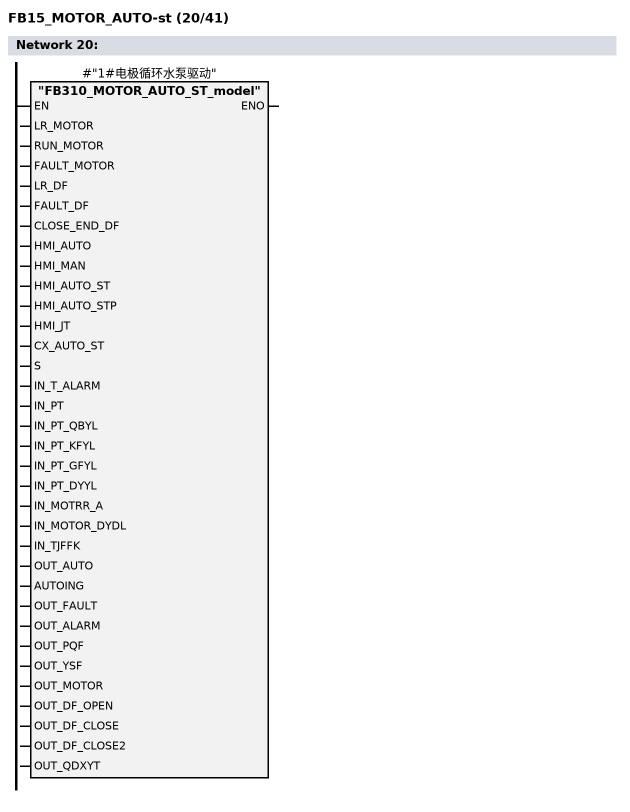
   RUNG wire#powerrail
      #"1#电极循环水泵驱动"(LR_MOTOR :=, RUN_MOTOR :=, FAULT_MOTOR :=, LR_DF :=, FAULT_DF :=, CLOSE_END_DF :=, HMI_AUTO :=, HMI_MAN :=, HMI_AUTO_ST :=, HMI_AUTO_STP :=, HMI_JT :=, CX_AUTO_ST :=, S :=, IN_T_ALARM :=, IN_PT :=, IN_PT_QBYL :=, IN_PT_KFYL :=, IN_PT_GFYL :=, IN_PT_DYYL :=, IN_MOTRR_A :=, IN_MOTOR_DYDL :=, IN_TJFFK :=, OUT_AUTO :=, AUTOING :=, OUT_FAULT :=, OUT_ALARM :=, OUT_PQF :=, OUT_YSF :=, OUT_MOTOR :=, OUT_DF_OPEN :=, OUT_DF_CLOSE :=, OUT_DF_CLOSE2 :=, OUT_QDXYT :=)
   END_RUNG
   // the same network as SCL:
   #"1#电极循环水泵驱动"();   // "FB310_MOTOR_AUTO_ST_model"
END_REGION

REGION Network 21
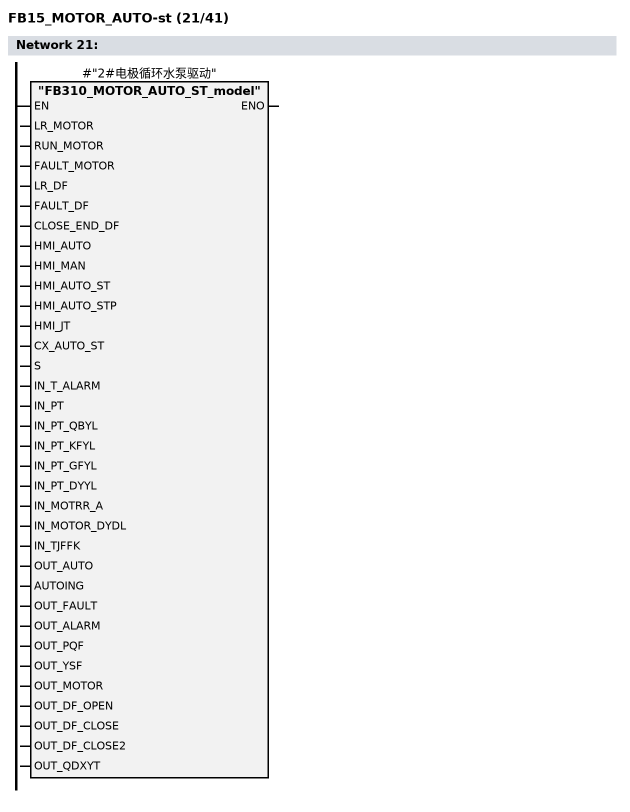
   RUNG wire#powerrail
      #"2#电极循环水泵驱动"(LR_MOTOR :=, RUN_MOTOR :=, FAULT_MOTOR :=, LR_DF :=, FAULT_DF :=, CLOSE_END_DF :=, HMI_AUTO :=, HMI_MAN :=, HMI_AUTO_ST :=, HMI_AUTO_STP :=, HMI_JT :=, CX_AUTO_ST :=, S :=, IN_T_ALARM :=, IN_PT :=, IN_PT_QBYL :=, IN_PT_KFYL :=, IN_PT_GFYL :=, IN_PT_DYYL :=, IN_MOTRR_A :=, IN_MOTOR_DYDL :=, IN_TJFFK :=, OUT_AUTO :=, AUTOING :=, OUT_FAULT :=, OUT_ALARM :=, OUT_PQF :=, OUT_YSF :=, OUT_MOTOR :=, OUT_DF_OPEN :=, OUT_DF_CLOSE :=, OUT_DF_CLOSE2 :=, OUT_QDXYT :=)
   END_RUNG
   // the same network as SCL:
   #"2#电极循环水泵驱动"();   // "FB310_MOTOR_AUTO_ST_model"
END_REGION

REGION Network 22
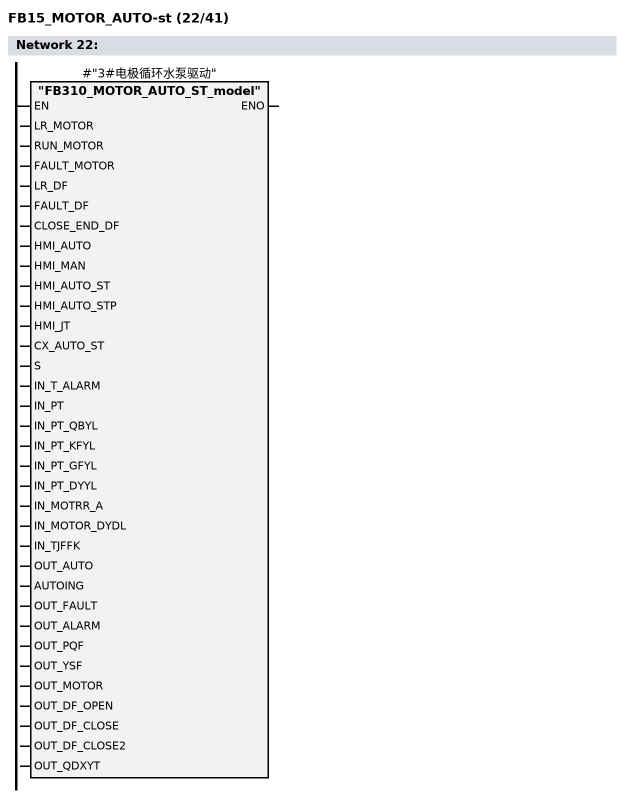
   RUNG wire#powerrail
      #"3#电极循环水泵驱动"(LR_MOTOR :=, RUN_MOTOR :=, FAULT_MOTOR :=, LR_DF :=, FAULT_DF :=, CLOSE_END_DF :=, HMI_AUTO :=, HMI_MAN :=, HMI_AUTO_ST :=, HMI_AUTO_STP :=, HMI_JT :=, CX_AUTO_ST :=, S :=, IN_T_ALARM :=, IN_PT :=, IN_PT_QBYL :=, IN_PT_KFYL :=, IN_PT_GFYL :=, IN_PT_DYYL :=, IN_MOTRR_A :=, IN_MOTOR_DYDL :=, IN_TJFFK :=, OUT_AUTO :=, AUTOING :=, OUT_FAULT :=, OUT_ALARM :=, OUT_PQF :=, OUT_YSF :=, OUT_MOTOR :=, OUT_DF_OPEN :=, OUT_DF_CLOSE :=, OUT_DF_CLOSE2 :=, OUT_QDXYT :=)
   END_RUNG
   // the same network as SCL:
   #"3#电极循环水泵驱动"();   // "FB310_MOTOR_AUTO_ST_model"
END_REGION

REGION Network 23
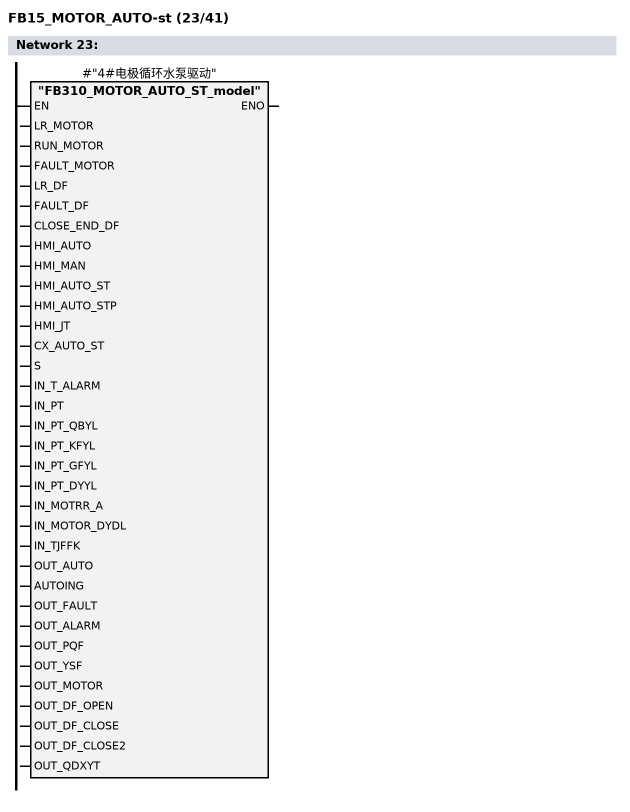
   RUNG wire#powerrail
      #"4#电极循环水泵驱动"(LR_MOTOR :=, RUN_MOTOR :=, FAULT_MOTOR :=, LR_DF :=, FAULT_DF :=, CLOSE_END_DF :=, HMI_AUTO :=, HMI_MAN :=, HMI_AUTO_ST :=, HMI_AUTO_STP :=, HMI_JT :=, CX_AUTO_ST :=, S :=, IN_T_ALARM :=, IN_PT :=, IN_PT_QBYL :=, IN_PT_KFYL :=, IN_PT_GFYL :=, IN_PT_DYYL :=, IN_MOTRR_A :=, IN_MOTOR_DYDL :=, IN_TJFFK :=, OUT_AUTO :=, AUTOING :=, OUT_FAULT :=, OUT_ALARM :=, OUT_PQF :=, OUT_YSF :=, OUT_MOTOR :=, OUT_DF_OPEN :=, OUT_DF_CLOSE :=, OUT_DF_CLOSE2 :=, OUT_QDXYT :=)
   END_RUNG
   // the same network as SCL:
   #"4#电极循环水泵驱动"();   // "FB310_MOTOR_AUTO_ST_model"
END_REGION

REGION Network 24
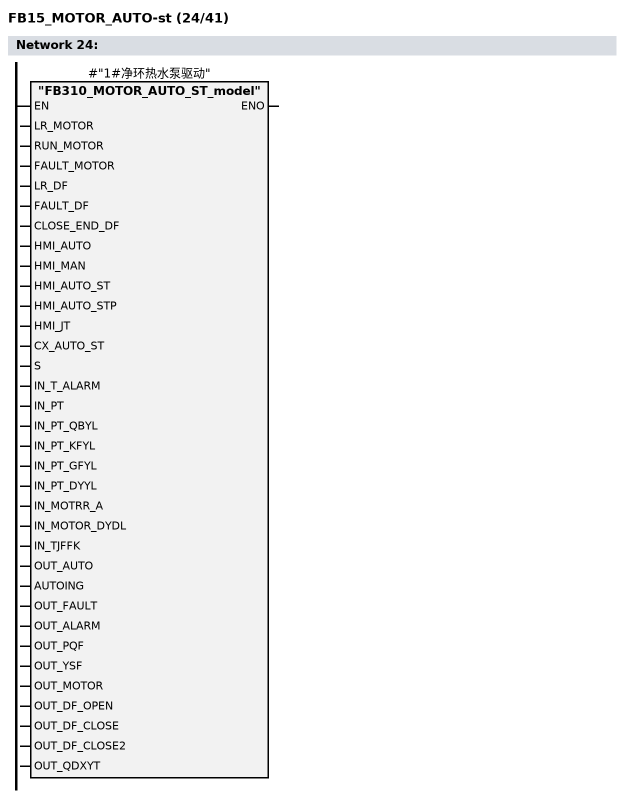
   RUNG wire#powerrail
      #"1#净环热水泵驱动"(LR_MOTOR :=, RUN_MOTOR :=, FAULT_MOTOR :=, LR_DF :=, FAULT_DF :=, CLOSE_END_DF :=, HMI_AUTO :=, HMI_MAN :=, HMI_AUTO_ST :=, HMI_AUTO_STP :=, HMI_JT :=, CX_AUTO_ST :=, S :=, IN_T_ALARM :=, IN_PT :=, IN_PT_QBYL :=, IN_PT_KFYL :=, IN_PT_GFYL :=, IN_PT_DYYL :=, IN_MOTRR_A :=, IN_MOTOR_DYDL :=, IN_TJFFK :=, OUT_AUTO :=, AUTOING :=, OUT_FAULT :=, OUT_ALARM :=, OUT_PQF :=, OUT_YSF :=, OUT_MOTOR :=, OUT_DF_OPEN :=, OUT_DF_CLOSE :=, OUT_DF_CLOSE2 :=, OUT_QDXYT :=)
   END_RUNG
   // the same network as SCL:
   #"1#净环热水泵驱动"();   // "FB310_MOTOR_AUTO_ST_model"
END_REGION

REGION Network 25
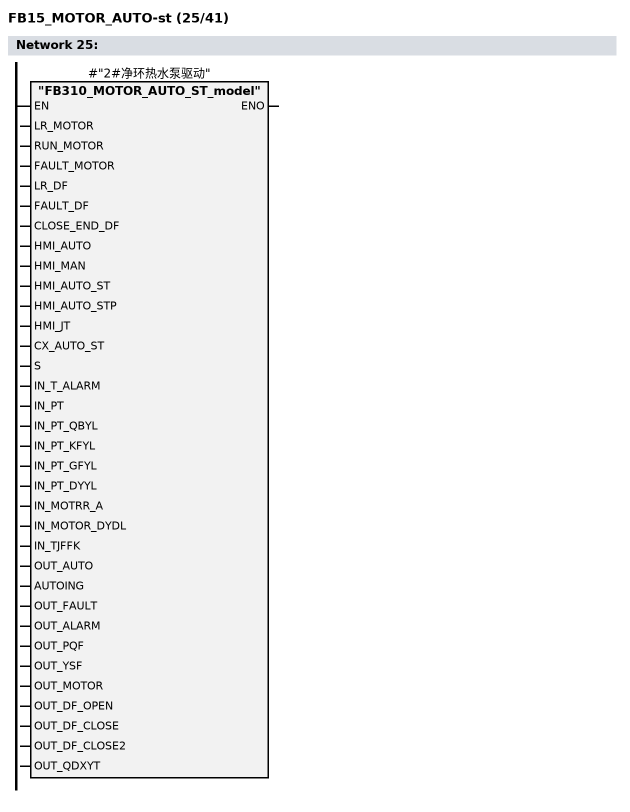
   RUNG wire#powerrail
      #"2#净环热水泵驱动"(LR_MOTOR :=, RUN_MOTOR :=, FAULT_MOTOR :=, LR_DF :=, FAULT_DF :=, CLOSE_END_DF :=, HMI_AUTO :=, HMI_MAN :=, HMI_AUTO_ST :=, HMI_AUTO_STP :=, HMI_JT :=, CX_AUTO_ST :=, S :=, IN_T_ALARM :=, IN_PT :=, IN_PT_QBYL :=, IN_PT_KFYL :=, IN_PT_GFYL :=, IN_PT_DYYL :=, IN_MOTRR_A :=, IN_MOTOR_DYDL :=, IN_TJFFK :=, OUT_AUTO :=, AUTOING :=, OUT_FAULT :=, OUT_ALARM :=, OUT_PQF :=, OUT_YSF :=, OUT_MOTOR :=, OUT_DF_OPEN :=, OUT_DF_CLOSE :=, OUT_DF_CLOSE2 :=, OUT_QDXYT :=)
   END_RUNG
   // the same network as SCL:
   #"2#净环热水泵驱动"();   // "FB310_MOTOR_AUTO_ST_model"
END_REGION

REGION Network 26
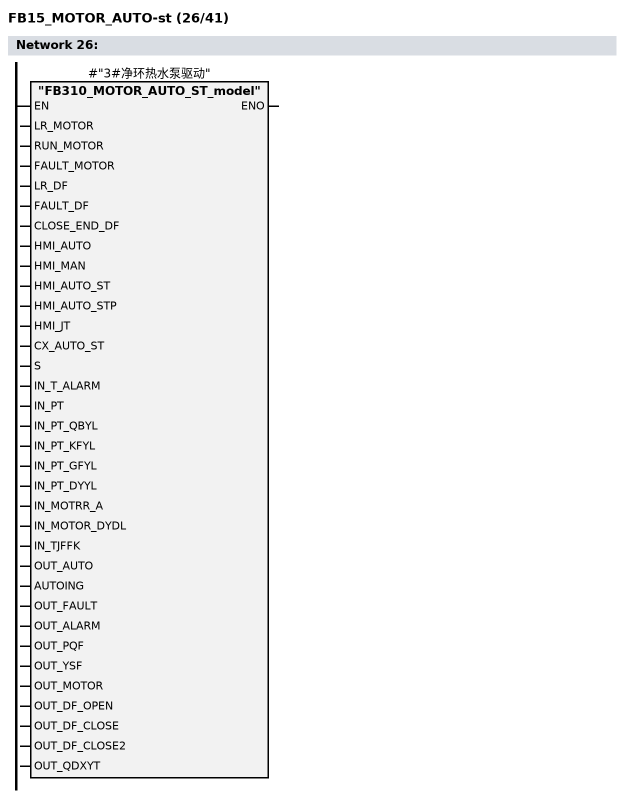
   RUNG wire#powerrail
      #"3#净环热水泵驱动"(LR_MOTOR :=, RUN_MOTOR :=, FAULT_MOTOR :=, LR_DF :=, FAULT_DF :=, CLOSE_END_DF :=, HMI_AUTO :=, HMI_MAN :=, HMI_AUTO_ST :=, HMI_AUTO_STP :=, HMI_JT :=, CX_AUTO_ST :=, S :=, IN_T_ALARM :=, IN_PT :=, IN_PT_QBYL :=, IN_PT_KFYL :=, IN_PT_GFYL :=, IN_PT_DYYL :=, IN_MOTRR_A :=, IN_MOTOR_DYDL :=, IN_TJFFK :=, OUT_AUTO :=, AUTOING :=, OUT_FAULT :=, OUT_ALARM :=, OUT_PQF :=, OUT_YSF :=, OUT_MOTOR :=, OUT_DF_OPEN :=, OUT_DF_CLOSE :=, OUT_DF_CLOSE2 :=, OUT_QDXYT :=)
   END_RUNG
   // the same network as SCL:
   #"3#净环热水泵驱动"();   // "FB310_MOTOR_AUTO_ST_model"
END_REGION

REGION Network 27
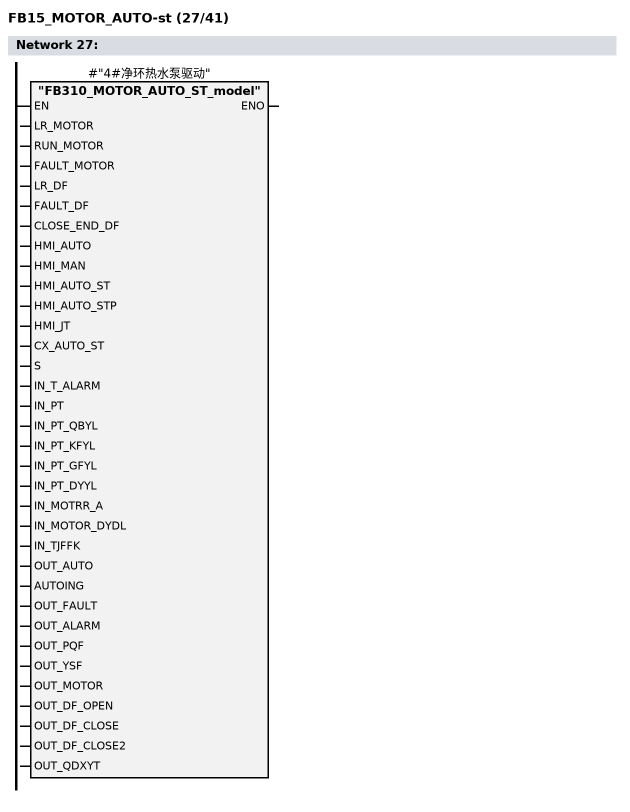
   RUNG wire#powerrail
      #"4#净环热水泵驱动"(LR_MOTOR :=, RUN_MOTOR :=, FAULT_MOTOR :=, LR_DF :=, FAULT_DF :=, CLOSE_END_DF :=, HMI_AUTO :=, HMI_MAN :=, HMI_AUTO_ST :=, HMI_AUTO_STP :=, HMI_JT :=, CX_AUTO_ST :=, S :=, IN_T_ALARM :=, IN_PT :=, IN_PT_QBYL :=, IN_PT_KFYL :=, IN_PT_GFYL :=, IN_PT_DYYL :=, IN_MOTRR_A :=, IN_MOTOR_DYDL :=, IN_TJFFK :=, OUT_AUTO :=, AUTOING :=, OUT_FAULT :=, OUT_ALARM :=, OUT_PQF :=, OUT_YSF :=, OUT_MOTOR :=, OUT_DF_OPEN :=, OUT_DF_CLOSE :=, OUT_DF_CLOSE2 :=, OUT_QDXYT :=)
   END_RUNG
   // the same network as SCL:
   #"4#净环热水泵驱动"();   // "FB310_MOTOR_AUTO_ST_model"
END_REGION

REGION Network 28
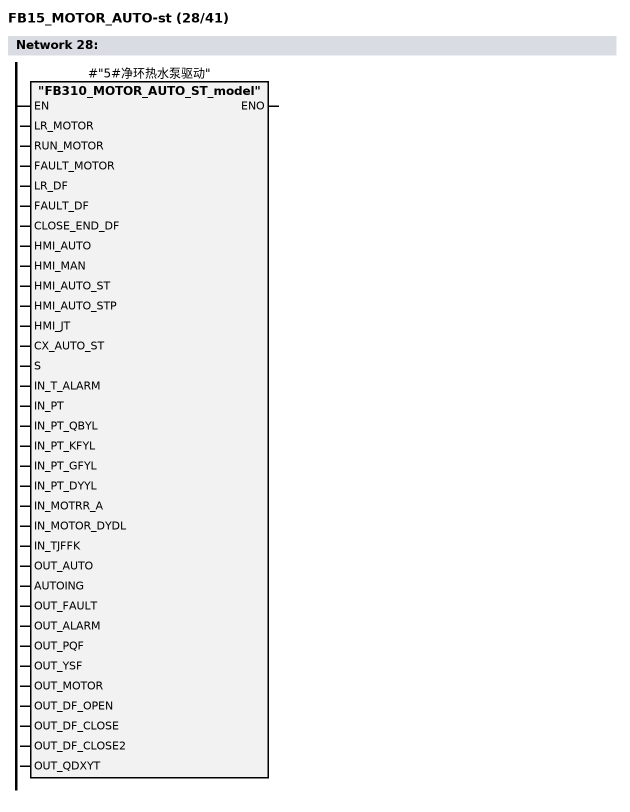
   RUNG wire#powerrail
      #"5#净环热水泵驱动"(LR_MOTOR :=, RUN_MOTOR :=, FAULT_MOTOR :=, LR_DF :=, FAULT_DF :=, CLOSE_END_DF :=, HMI_AUTO :=, HMI_MAN :=, HMI_AUTO_ST :=, HMI_AUTO_STP :=, HMI_JT :=, CX_AUTO_ST :=, S :=, IN_T_ALARM :=, IN_PT :=, IN_PT_QBYL :=, IN_PT_KFYL :=, IN_PT_GFYL :=, IN_PT_DYYL :=, IN_MOTRR_A :=, IN_MOTOR_DYDL :=, IN_TJFFK :=, OUT_AUTO :=, AUTOING :=, OUT_FAULT :=, OUT_ALARM :=, OUT_PQF :=, OUT_YSF :=, OUT_MOTOR :=, OUT_DF_OPEN :=, OUT_DF_CLOSE :=, OUT_DF_CLOSE2 :=, OUT_QDXYT :=)
   END_RUNG
   // the same network as SCL:
   #"5#净环热水泵驱动"();   // "FB310_MOTOR_AUTO_ST_model"
END_REGION

REGION Network 29
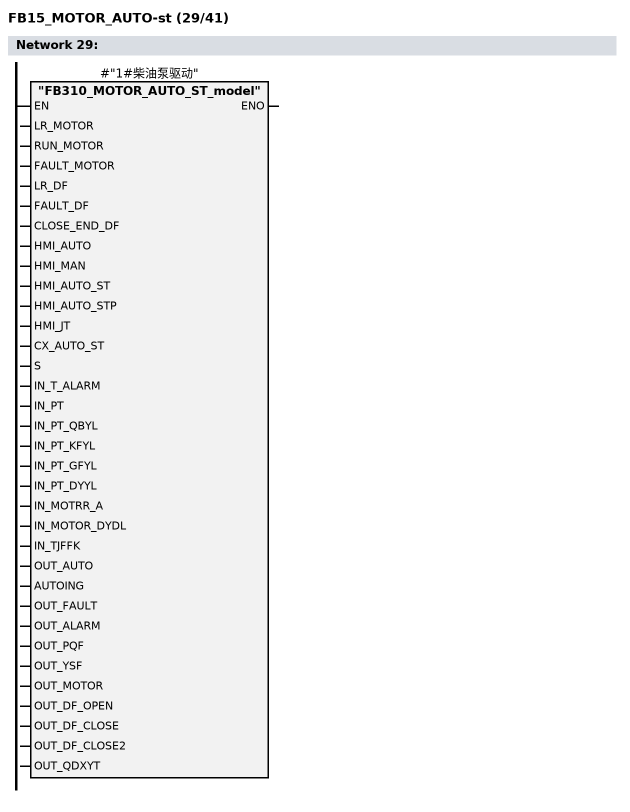
   RUNG wire#powerrail
      #"1#柴油泵驱动"(LR_MOTOR :=, RUN_MOTOR :=, FAULT_MOTOR :=, LR_DF :=, FAULT_DF :=, CLOSE_END_DF :=, HMI_AUTO :=, HMI_MAN :=, HMI_AUTO_ST :=, HMI_AUTO_STP :=, HMI_JT :=, CX_AUTO_ST :=, S :=, IN_T_ALARM :=, IN_PT :=, IN_PT_QBYL :=, IN_PT_KFYL :=, IN_PT_GFYL :=, IN_PT_DYYL :=, IN_MOTRR_A :=, IN_MOTOR_DYDL :=, IN_TJFFK :=, OUT_AUTO :=, AUTOING :=, OUT_FAULT :=, OUT_ALARM :=, OUT_PQF :=, OUT_YSF :=, OUT_MOTOR :=, OUT_DF_OPEN :=, OUT_DF_CLOSE :=, OUT_DF_CLOSE2 :=, OUT_QDXYT :=)
   END_RUNG
   // the same network as SCL:
   #"1#柴油泵驱动"();   // "FB310_MOTOR_AUTO_ST_model"
END_REGION

REGION Network 30
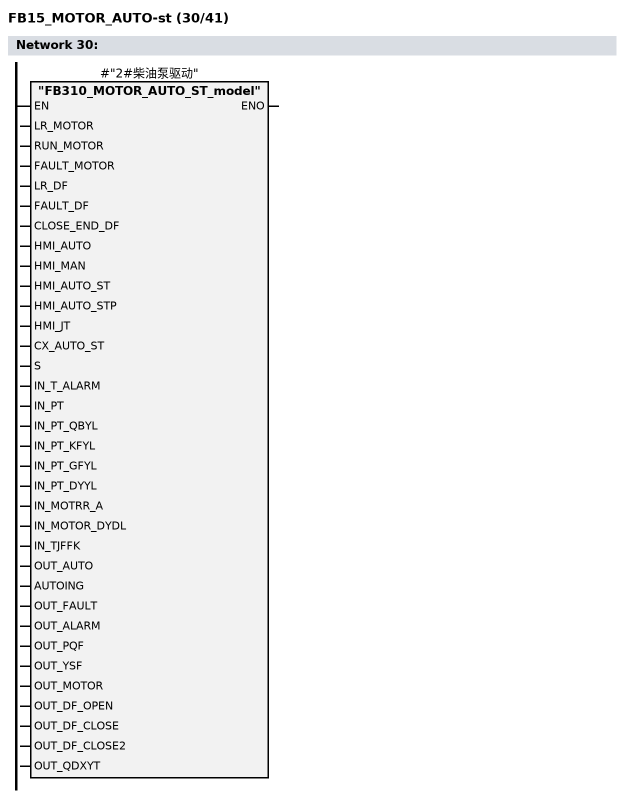
   RUNG wire#powerrail
      #"2#柴油泵驱动"(LR_MOTOR :=, RUN_MOTOR :=, FAULT_MOTOR :=, LR_DF :=, FAULT_DF :=, CLOSE_END_DF :=, HMI_AUTO :=, HMI_MAN :=, HMI_AUTO_ST :=, HMI_AUTO_STP :=, HMI_JT :=, CX_AUTO_ST :=, S :=, IN_T_ALARM :=, IN_PT :=, IN_PT_QBYL :=, IN_PT_KFYL :=, IN_PT_GFYL :=, IN_PT_DYYL :=, IN_MOTRR_A :=, IN_MOTOR_DYDL :=, IN_TJFFK :=, OUT_AUTO :=, AUTOING :=, OUT_FAULT :=, OUT_ALARM :=, OUT_PQF :=, OUT_YSF :=, OUT_MOTOR :=, OUT_DF_OPEN :=, OUT_DF_CLOSE :=, OUT_DF_CLOSE2 :=, OUT_QDXYT :=)
   END_RUNG
   // the same network as SCL:
   #"2#柴油泵驱动"();   // "FB310_MOTOR_AUTO_ST_model"
END_REGION

REGION Network 31
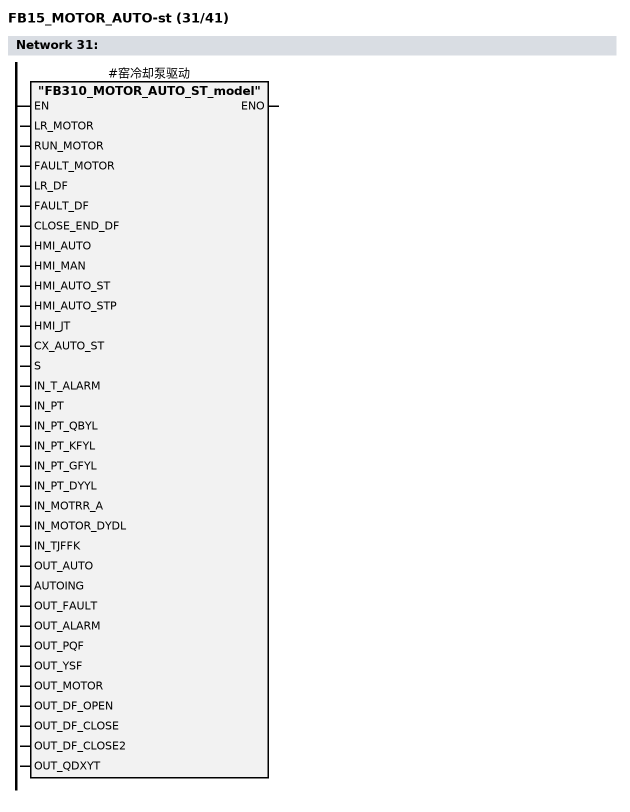
   RUNG wire#powerrail
      #窑冷却泵驱动(LR_MOTOR :=, RUN_MOTOR :=, FAULT_MOTOR :=, LR_DF :=, FAULT_DF :=, CLOSE_END_DF :=, HMI_AUTO :=, HMI_MAN :=, HMI_AUTO_ST :=, HMI_AUTO_STP :=, HMI_JT :=, CX_AUTO_ST :=, S :=, IN_T_ALARM :=, IN_PT :=, IN_PT_QBYL :=, IN_PT_KFYL :=, IN_PT_GFYL :=, IN_PT_DYYL :=, IN_MOTRR_A :=, IN_MOTOR_DYDL :=, IN_TJFFK :=, OUT_AUTO :=, AUTOING :=, OUT_FAULT :=, OUT_ALARM :=, OUT_PQF :=, OUT_YSF :=, OUT_MOTOR :=, OUT_DF_OPEN :=, OUT_DF_CLOSE :=, OUT_DF_CLOSE2 :=, OUT_QDXYT :=)
   END_RUNG
   // the same network as SCL:
   #窑冷却泵驱动();   // "FB310_MOTOR_AUTO_ST_model"
END_REGION

REGION Network 32
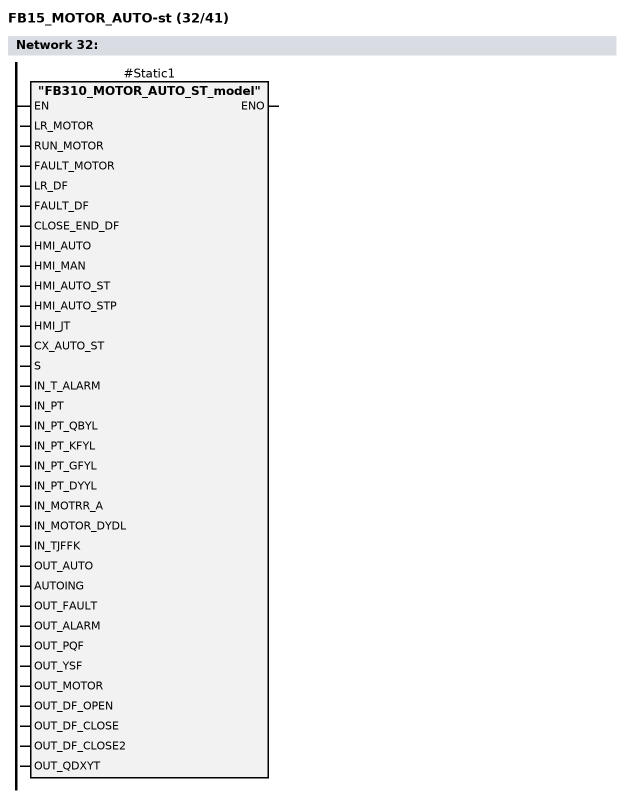
   RUNG wire#powerrail
      #Static1(LR_MOTOR :=, RUN_MOTOR :=, FAULT_MOTOR :=, LR_DF :=, FAULT_DF :=, CLOSE_END_DF :=, HMI_AUTO :=, HMI_MAN :=, HMI_AUTO_ST :=, HMI_AUTO_STP :=, HMI_JT :=, CX_AUTO_ST :=, S :=, IN_T_ALARM :=, IN_PT :=, IN_PT_QBYL :=, IN_PT_KFYL :=, IN_PT_GFYL :=, IN_PT_DYYL :=, IN_MOTRR_A :=, IN_MOTOR_DYDL :=, IN_TJFFK :=, OUT_AUTO :=, AUTOING :=, OUT_FAULT :=, OUT_ALARM :=, OUT_PQF :=, OUT_YSF :=, OUT_MOTOR :=, OUT_DF_OPEN :=, OUT_DF_CLOSE :=, OUT_DF_CLOSE2 :=, OUT_QDXYT :=)
   END_RUNG
   // the same network as SCL:
   #Static1();   // "FB310_MOTOR_AUTO_ST_model"
END_REGION

REGION Network 33
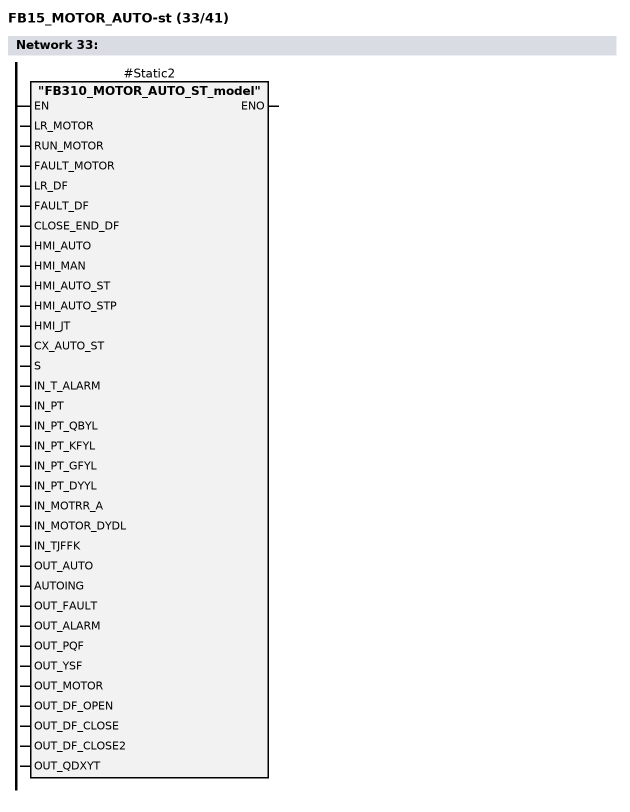
   RUNG wire#powerrail
      #Static2(LR_MOTOR :=, RUN_MOTOR :=, FAULT_MOTOR :=, LR_DF :=, FAULT_DF :=, CLOSE_END_DF :=, HMI_AUTO :=, HMI_MAN :=, HMI_AUTO_ST :=, HMI_AUTO_STP :=, HMI_JT :=, CX_AUTO_ST :=, S :=, IN_T_ALARM :=, IN_PT :=, IN_PT_QBYL :=, IN_PT_KFYL :=, IN_PT_GFYL :=, IN_PT_DYYL :=, IN_MOTRR_A :=, IN_MOTOR_DYDL :=, IN_TJFFK :=, OUT_AUTO :=, AUTOING :=, OUT_FAULT :=, OUT_ALARM :=, OUT_PQF :=, OUT_YSF :=, OUT_MOTOR :=, OUT_DF_OPEN :=, OUT_DF_CLOSE :=, OUT_DF_CLOSE2 :=, OUT_QDXYT :=)
   END_RUNG
   // the same network as SCL:
   #Static2();   // "FB310_MOTOR_AUTO_ST_model"
END_REGION

REGION Network 34
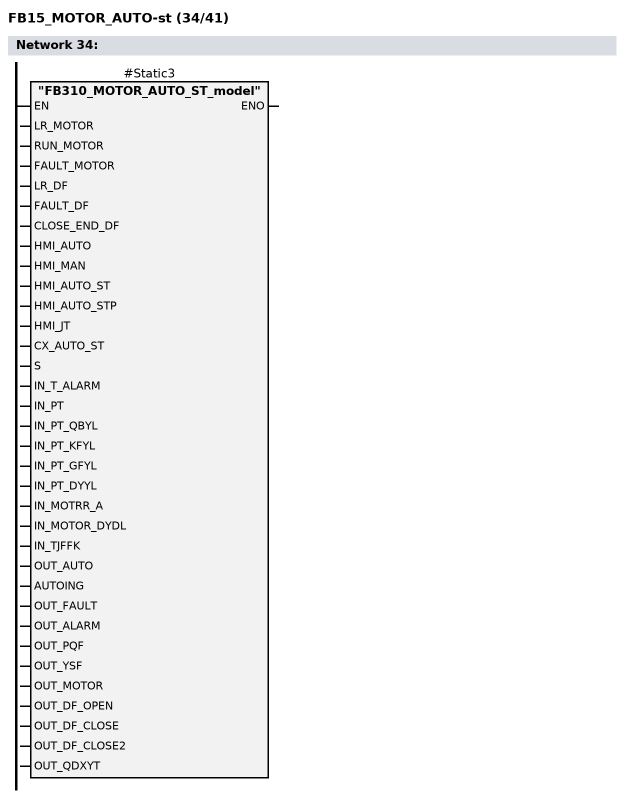
   RUNG wire#powerrail
      #Static3(LR_MOTOR :=, RUN_MOTOR :=, FAULT_MOTOR :=, LR_DF :=, FAULT_DF :=, CLOSE_END_DF :=, HMI_AUTO :=, HMI_MAN :=, HMI_AUTO_ST :=, HMI_AUTO_STP :=, HMI_JT :=, CX_AUTO_ST :=, S :=, IN_T_ALARM :=, IN_PT :=, IN_PT_QBYL :=, IN_PT_KFYL :=, IN_PT_GFYL :=, IN_PT_DYYL :=, IN_MOTRR_A :=, IN_MOTOR_DYDL :=, IN_TJFFK :=, OUT_AUTO :=, AUTOING :=, OUT_FAULT :=, OUT_ALARM :=, OUT_PQF :=, OUT_YSF :=, OUT_MOTOR :=, OUT_DF_OPEN :=, OUT_DF_CLOSE :=, OUT_DF_CLOSE2 :=, OUT_QDXYT :=)
   END_RUNG
   // the same network as SCL:
   #Static3();   // "FB310_MOTOR_AUTO_ST_model"
END_REGION

REGION Network 35
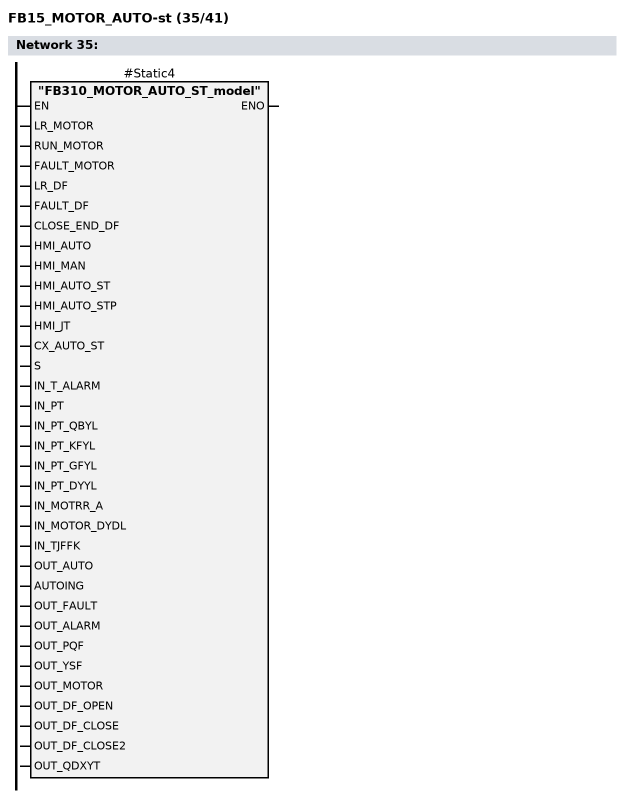
   RUNG wire#powerrail
      #Static4(LR_MOTOR :=, RUN_MOTOR :=, FAULT_MOTOR :=, LR_DF :=, FAULT_DF :=, CLOSE_END_DF :=, HMI_AUTO :=, HMI_MAN :=, HMI_AUTO_ST :=, HMI_AUTO_STP :=, HMI_JT :=, CX_AUTO_ST :=, S :=, IN_T_ALARM :=, IN_PT :=, IN_PT_QBYL :=, IN_PT_KFYL :=, IN_PT_GFYL :=, IN_PT_DYYL :=, IN_MOTRR_A :=, IN_MOTOR_DYDL :=, IN_TJFFK :=, OUT_AUTO :=, AUTOING :=, OUT_FAULT :=, OUT_ALARM :=, OUT_PQF :=, OUT_YSF :=, OUT_MOTOR :=, OUT_DF_OPEN :=, OUT_DF_CLOSE :=, OUT_DF_CLOSE2 :=, OUT_QDXYT :=)
   END_RUNG
   // the same network as SCL:
   #Static4();   // "FB310_MOTOR_AUTO_ST_model"
END_REGION

REGION Network 36
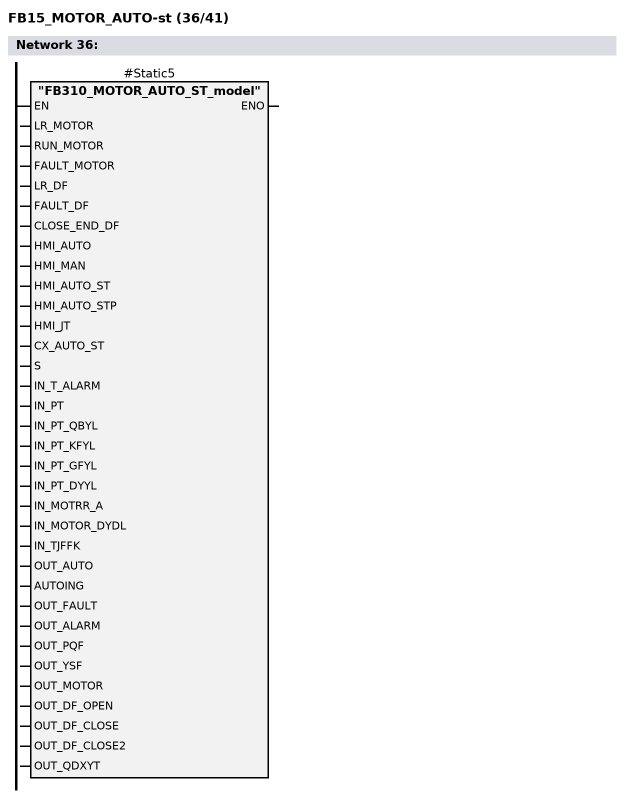
   RUNG wire#powerrail
      #Static5(LR_MOTOR :=, RUN_MOTOR :=, FAULT_MOTOR :=, LR_DF :=, FAULT_DF :=, CLOSE_END_DF :=, HMI_AUTO :=, HMI_MAN :=, HMI_AUTO_ST :=, HMI_AUTO_STP :=, HMI_JT :=, CX_AUTO_ST :=, S :=, IN_T_ALARM :=, IN_PT :=, IN_PT_QBYL :=, IN_PT_KFYL :=, IN_PT_GFYL :=, IN_PT_DYYL :=, IN_MOTRR_A :=, IN_MOTOR_DYDL :=, IN_TJFFK :=, OUT_AUTO :=, AUTOING :=, OUT_FAULT :=, OUT_ALARM :=, OUT_PQF :=, OUT_YSF :=, OUT_MOTOR :=, OUT_DF_OPEN :=, OUT_DF_CLOSE :=, OUT_DF_CLOSE2 :=, OUT_QDXYT :=)
   END_RUNG
   // the same network as SCL:
   #Static5();   // "FB310_MOTOR_AUTO_ST_model"
END_REGION

REGION Network 37
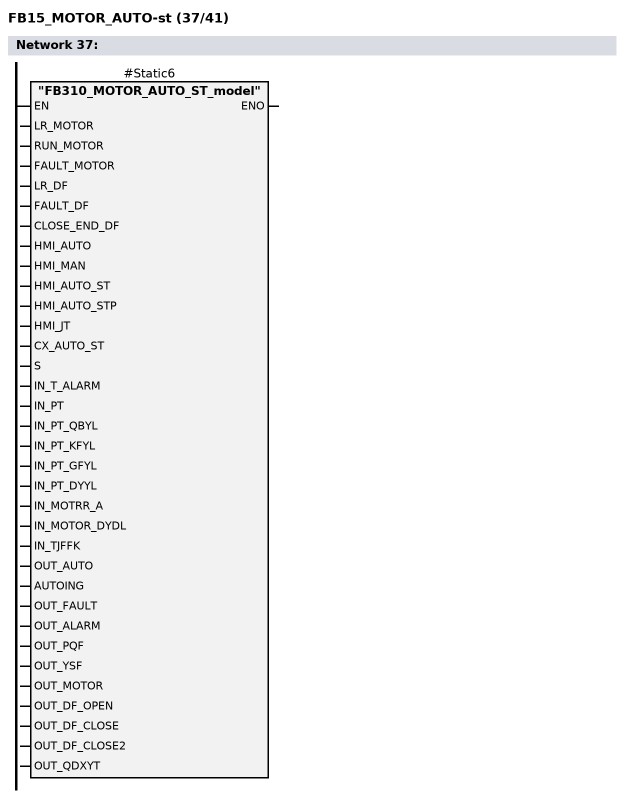
   RUNG wire#powerrail
      #Static6(LR_MOTOR :=, RUN_MOTOR :=, FAULT_MOTOR :=, LR_DF :=, FAULT_DF :=, CLOSE_END_DF :=, HMI_AUTO :=, HMI_MAN :=, HMI_AUTO_ST :=, HMI_AUTO_STP :=, HMI_JT :=, CX_AUTO_ST :=, S :=, IN_T_ALARM :=, IN_PT :=, IN_PT_QBYL :=, IN_PT_KFYL :=, IN_PT_GFYL :=, IN_PT_DYYL :=, IN_MOTRR_A :=, IN_MOTOR_DYDL :=, IN_TJFFK :=, OUT_AUTO :=, AUTOING :=, OUT_FAULT :=, OUT_ALARM :=, OUT_PQF :=, OUT_YSF :=, OUT_MOTOR :=, OUT_DF_OPEN :=, OUT_DF_CLOSE :=, OUT_DF_CLOSE2 :=, OUT_QDXYT :=)
   END_RUNG
   // the same network as SCL:
   #Static6();   // "FB310_MOTOR_AUTO_ST_model"
END_REGION

REGION Network 38
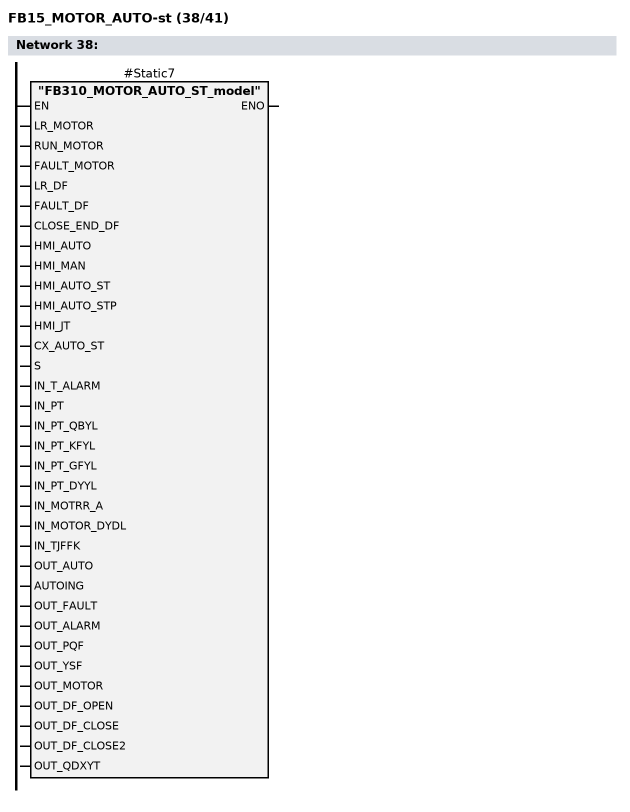
   RUNG wire#powerrail
      #Static7(LR_MOTOR :=, RUN_MOTOR :=, FAULT_MOTOR :=, LR_DF :=, FAULT_DF :=, CLOSE_END_DF :=, HMI_AUTO :=, HMI_MAN :=, HMI_AUTO_ST :=, HMI_AUTO_STP :=, HMI_JT :=, CX_AUTO_ST :=, S :=, IN_T_ALARM :=, IN_PT :=, IN_PT_QBYL :=, IN_PT_KFYL :=, IN_PT_GFYL :=, IN_PT_DYYL :=, IN_MOTRR_A :=, IN_MOTOR_DYDL :=, IN_TJFFK :=, OUT_AUTO :=, AUTOING :=, OUT_FAULT :=, OUT_ALARM :=, OUT_PQF :=, OUT_YSF :=, OUT_MOTOR :=, OUT_DF_OPEN :=, OUT_DF_CLOSE :=, OUT_DF_CLOSE2 :=, OUT_QDXYT :=)
   END_RUNG
   // the same network as SCL:
   #Static7();   // "FB310_MOTOR_AUTO_ST_model"
END_REGION

REGION Network 39
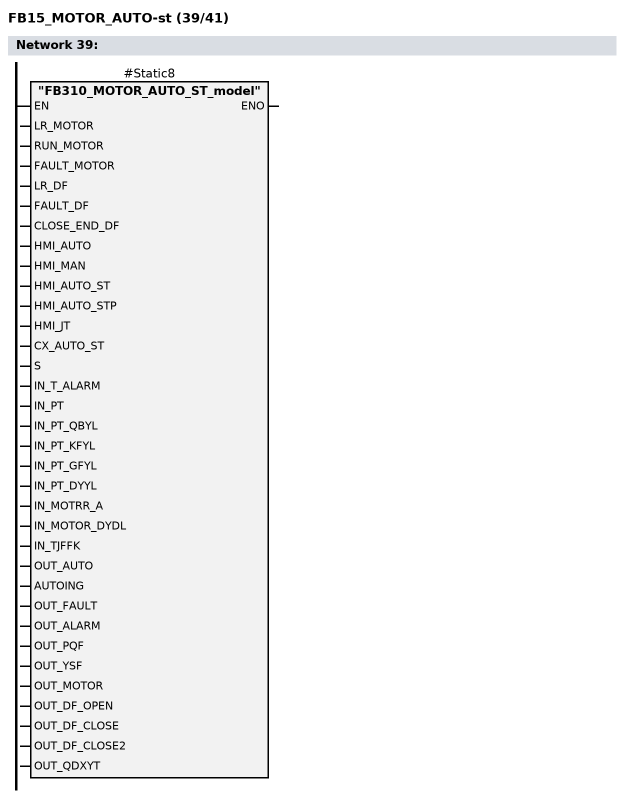
   RUNG wire#powerrail
      #Static8(LR_MOTOR :=, RUN_MOTOR :=, FAULT_MOTOR :=, LR_DF :=, FAULT_DF :=, CLOSE_END_DF :=, HMI_AUTO :=, HMI_MAN :=, HMI_AUTO_ST :=, HMI_AUTO_STP :=, HMI_JT :=, CX_AUTO_ST :=, S :=, IN_T_ALARM :=, IN_PT :=, IN_PT_QBYL :=, IN_PT_KFYL :=, IN_PT_GFYL :=, IN_PT_DYYL :=, IN_MOTRR_A :=, IN_MOTOR_DYDL :=, IN_TJFFK :=, OUT_AUTO :=, AUTOING :=, OUT_FAULT :=, OUT_ALARM :=, OUT_PQF :=, OUT_YSF :=, OUT_MOTOR :=, OUT_DF_OPEN :=, OUT_DF_CLOSE :=, OUT_DF_CLOSE2 :=, OUT_QDXYT :=)
   END_RUNG
   // the same network as SCL:
   #Static8();   // "FB310_MOTOR_AUTO_ST_model"
END_REGION

REGION Network 40
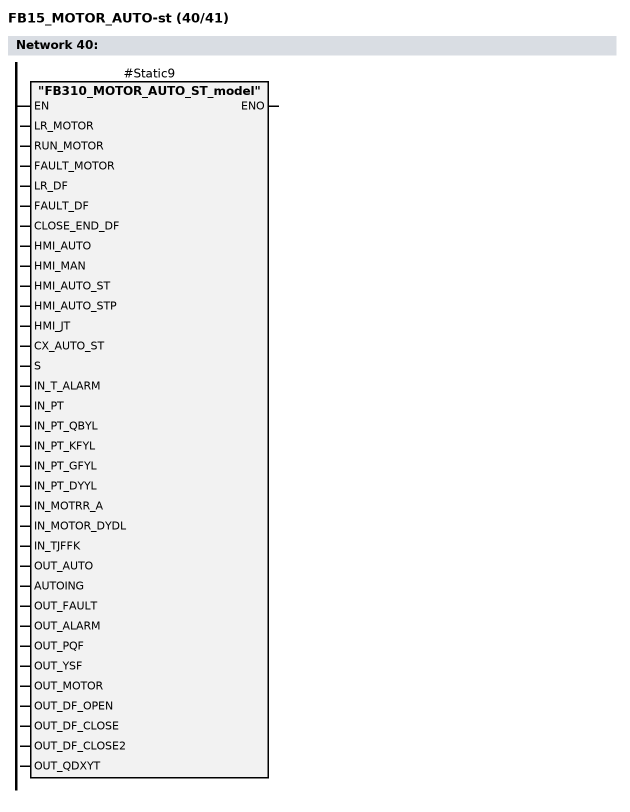
   RUNG wire#powerrail
      #Static9(LR_MOTOR :=, RUN_MOTOR :=, FAULT_MOTOR :=, LR_DF :=, FAULT_DF :=, CLOSE_END_DF :=, HMI_AUTO :=, HMI_MAN :=, HMI_AUTO_ST :=, HMI_AUTO_STP :=, HMI_JT :=, CX_AUTO_ST :=, S :=, IN_T_ALARM :=, IN_PT :=, IN_PT_QBYL :=, IN_PT_KFYL :=, IN_PT_GFYL :=, IN_PT_DYYL :=, IN_MOTRR_A :=, IN_MOTOR_DYDL :=, IN_TJFFK :=, OUT_AUTO :=, AUTOING :=, OUT_FAULT :=, OUT_ALARM :=, OUT_PQF :=, OUT_YSF :=, OUT_MOTOR :=, OUT_DF_OPEN :=, OUT_DF_CLOSE :=, OUT_DF_CLOSE2 :=, OUT_QDXYT :=)
   END_RUNG
   // the same network as SCL:
   #Static9();   // "FB310_MOTOR_AUTO_ST_model"
END_REGION

REGION Network 41
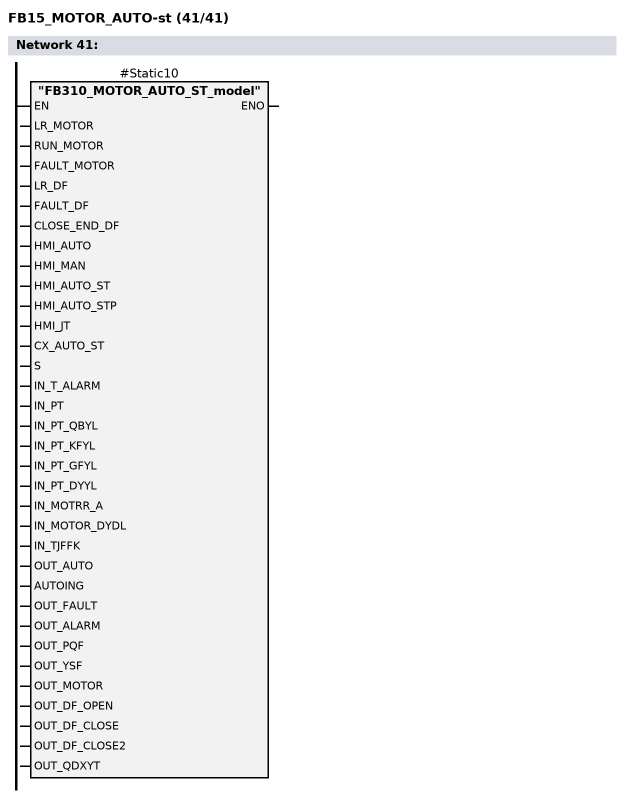
   RUNG wire#powerrail
      #Static10(LR_MOTOR :=, RUN_MOTOR :=, FAULT_MOTOR :=, LR_DF :=, FAULT_DF :=, CLOSE_END_DF :=, HMI_AUTO :=, HMI_MAN :=, HMI_AUTO_ST :=, HMI_AUTO_STP :=, HMI_JT :=, CX_AUTO_ST :=, S :=, IN_T_ALARM :=, IN_PT :=, IN_PT_QBYL :=, IN_PT_KFYL :=, IN_PT_GFYL :=, IN_PT_DYYL :=, IN_MOTRR_A :=, IN_MOTOR_DYDL :=, IN_TJFFK :=, OUT_AUTO :=, AUTOING :=, OUT_FAULT :=, OUT_ALARM :=, OUT_PQF :=, OUT_YSF :=, OUT_MOTOR :=, OUT_DF_OPEN :=, OUT_DF_CLOSE :=, OUT_DF_CLOSE2 :=, OUT_QDXYT :=)
   END_RUNG
   // the same network as SCL:
   #Static10();   // "FB310_MOTOR_AUTO_ST_model"
END_REGION
END_FUNCTION_BLOCK

FUNCTION_BLOCK "电机_冷却塔风机"   // FB301, LAD
{ S7_Optimized_Access := 'FALSE' }
VERSION : 0.1
// 用于电机的启停控制。具有手动/自动模式，手动模式通过画面的启停按钮启动；自动根据外部的启停条件启动。
// 故障判断：有输出无运行反馈信号持续x秒报价；热过载跳脱报警。
// 有单次运行时间和累计运行时间计时和复位。
   VAR_INPUT
      LR : Bool;
      READY : Bool;
      RUN : Bool;
      FAULT : Bool;
      HMI_ST : Bool;
      HMI_STP : Bool;
      MA : Bool;
      AUTO : Bool;
      FLT_RST : Bool;
      TIME_EN : Bool := TRUE;
      TIME_RST : Bool;
      JT : Bool;
      S : Bool;
      TIME_FAULT : Time := T#120S;
   END_VAR
   VAR_OUTPUT
      TIME_RUN : Real;   // 单次运行时间
      TIME_ALL : Real;   // 累加运行时间
   END_VAR
   VAR_IN_OUT
      OUT : Bool;
      FAULT_STOP : Bool;
   END_VAR
   VAR
      MAN_OUT : Bool;
      P1 : Bool;
      P2 : Bool;
      T_FAULT1 : IEC_TIMER;
      T_FAULT2 : IEC_TIMER;
      STAT1 : Real;   // 单次运行时间
      STAT2 : Real;   // 累计运行时间
   END_VAR
   VAR_TEMP   // added for the SCL form of the ladder/FBD networks
      _w1 : Bool;
      _w2 : Bool;
   END_VAR
BEGIN

REGION Network 1
   // 手动输出
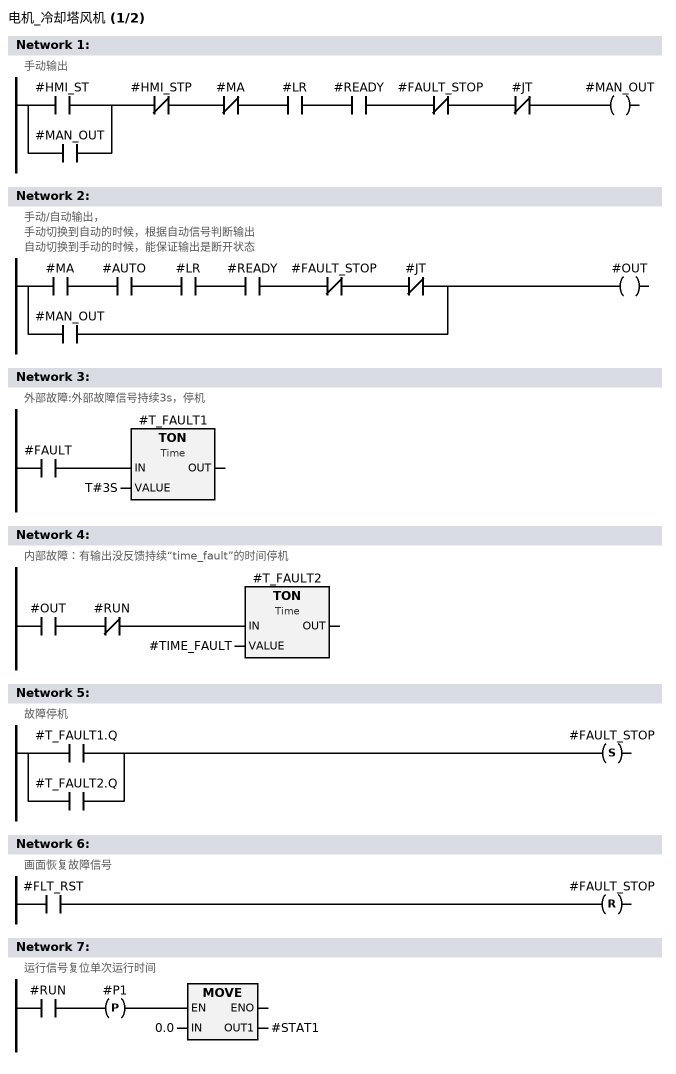
   RUNG wire#powerrail
      Contact( #HMI_ST )
      wire#w1
      I_Contact( #HMI_STP )
      I_Contact( #MA )
      Contact( #LR )
      Contact( #READY )
      I_Contact( #FAULT_STOP )
      I_Contact( #JT )
      Coil( #MAN_OUT )
   END_RUNG
   RUNG wire#powerrail
      Contact( #MAN_OUT )
   END_RUNG wire#w1
   // the same network as SCL:
   #MAN_OUT := (#HMI_ST OR #MAN_OUT) AND NOT #HMI_STP AND NOT #MA AND #LR AND #READY AND NOT #FAULT_STOP AND NOT #JT;
END_REGION

REGION Network 2
   // 手动/自动输出，
   // 手动切换到自动的时候，根据自动信号判断输出
   // 自动切换到手动的时候，能保证输出是断开状态
   RUNG wire#powerrail
      Contact( #MA )
      Contact( #AUTO )
      Contact( #LR )
      Contact( #READY )
      I_Contact( #FAULT_STOP )
      I_Contact( #JT )
      wire#w1
      Coil( #OUT )
   END_RUNG
   RUNG wire#powerrail
      Contact( #MAN_OUT )
   END_RUNG wire#w1
   // the same network as SCL:
   #OUT := (#MA AND #AUTO AND #LR AND #READY AND NOT #FAULT_STOP AND NOT #JT) OR #MAN_OUT;
END_REGION

REGION Network 3
   // 外部故障:外部故障信号持续3s，停机
   #T_FAULT1.TON(IN := #FAULT, PT := T#3S);   // TON coil
END_REGION

REGION Network 4
   // 内部故障：有输出没反馈持续“time_fault”的时间停机
   #T_FAULT2.TON(IN := #OUT AND NOT #RUN, PT := #TIME_FAULT);   // TON coil
END_REGION

REGION Network 5
   // 故障停机
   RUNG wire#powerrail
      Contact( #T_FAULT1.Q )
      wire#w1
      S_Coil( #FAULT_STOP )
   END_RUNG
   RUNG wire#powerrail
      Contact( #T_FAULT2.Q )
   END_RUNG wire#w1
   // the same network as SCL:
   IF #T_FAULT1.Q OR #T_FAULT2.Q THEN #FAULT_STOP := TRUE; END_IF;
END_REGION

REGION Network 6
   // 画面恢复故障信号
   RUNG wire#powerrail
      Contact( #FLT_RST )
      R_Coil( #FAULT_STOP )
   END_RUNG
   // the same network as SCL:
   IF #FLT_RST THEN #FAULT_STOP := FALSE; END_IF;
END_REGION

REGION Network 7
   // 运行信号复位单次运行时间
   RUNG wire#powerrail
      Contact( #RUN )
      P_Trig( #P1 )
      Move(in := 0.0, out1 => #STAT1)
   END_RUNG
   // the same network as SCL:
   #_w1 := #RUN AND NOT #P1;   // rising edge
   #P1 := #RUN;
   IF #_w1 THEN #STAT1 := 0.0; END_IF;
END_REGION

REGION Network 8
   // 有运行信号无故障信号则开始累加 单次运行时间和累计运行时间
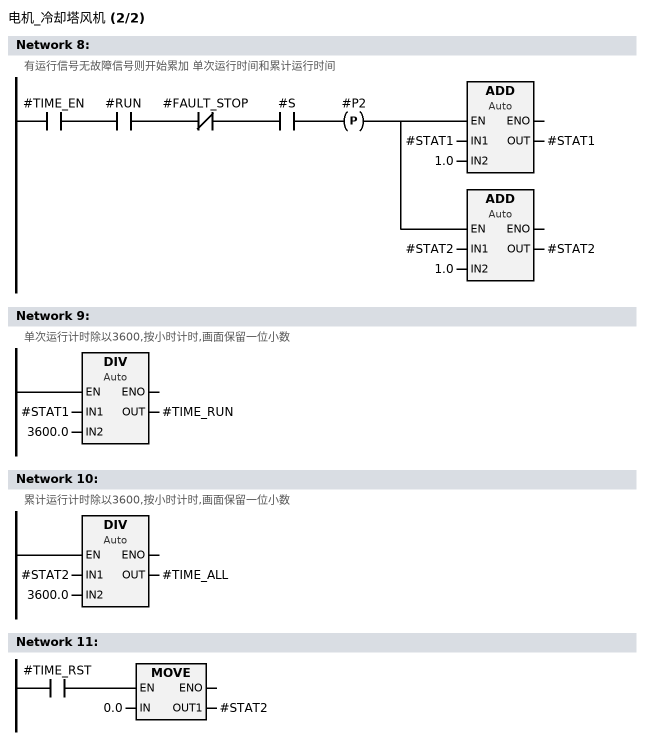
   RUNG wire#powerrail
      Contact( #TIME_EN )
      Contact( #RUN )
      I_Contact( #FAULT_STOP )
      Contact( #S )
      P_Trig( #P2 )
      wire#w1
      Add(in1 := #STAT1, in2 := 1.0, out => #STAT1)
   END_RUNG
   RUNG wire#w1
      Add(in1 := #STAT2, in2 := 1.0, out => #STAT2)
   END_RUNG
   // the same network as SCL:
   #_w1 := #TIME_EN AND #RUN AND NOT #FAULT_STOP AND #S;
   #_w2 := #_w1 AND NOT #P2;   // rising edge
   #P2 := #_w1;
   IF #_w2 THEN
       #STAT1 := #STAT1 + 1.0;
       #STAT2 := #STAT2 + 1.0;
   END_IF;
END_REGION

REGION Network 9
   // 单次运行计时除以3600,按小时计时,画面保留一位小数
   RUNG wire#powerrail
      Div(in1 := #STAT1, in2 := 3600.0, out => #TIME_RUN)
   END_RUNG
   // the same network as SCL:
   #TIME_RUN := #STAT1 / 3600.0;
END_REGION

REGION Network 10
   // 累计运行计时除以3600,按小时计时,画面保留一位小数
   RUNG wire#powerrail
      Div(in1 := #STAT2, in2 := 3600.0, out => #TIME_ALL)
   END_RUNG
   // the same network as SCL:
   #TIME_ALL := #STAT2 / 3600.0;
END_REGION

REGION Network 11
   RUNG wire#powerrail
      Contact( #TIME_RST )
      Move(in := 0.0, out1 => #STAT2)
   END_RUNG
   // the same network as SCL:
   IF #TIME_RST THEN #STAT2 := 0.0; END_IF;
END_REGION
END_FUNCTION_BLOCK

FUNCTION_BLOCK "阀门_MODEL"   // FB302, LAD
{ S7_Optimized_Access := 'FALSE' }
VERSION : 0.1
   VAR_INPUT
      READY : Bool;
      RUN : Bool;
      FAULT : Bool;
      OPEN_END : Bool;
      CLOSE_END : Bool;
      HMI_OPEN : Bool;
      HMI_CLOSE : Bool;
      MA : Bool;
      AUTO_OPEN : Bool;
      AUTO_CLOSE : Bool;
   END_VAR
   VAR_IN_OUT
      QD_OPEN : Bool;
      QD_CLOSE : Bool;
   END_VAR
BEGIN

REGION Network 1
